   	OWF_Key[313,9]:=1836248757;
   	OWF_Key[313,10]:=799041735;
   	OWF_Key[313,11]:=206920278;
   	OWF_Key[313,12]:=1670185075;
   	OWF_Key[314,0]:=167288513;
   	OWF_Key[314,1]:=1823765264;
   	OWF_Key[314,2]:=1024405687;
   	OWF_Key[314,3]:=1305159346;
   	OWF_Key[314,4]:=1207657799;
   	OWF_Key[314,5]:=1657238232;
   	OWF_Key[314,6]:=1138840138;
   	OWF_Key[314,7]:=1308155371;
   	OWF_Key[314,8]:=444304420;
   	OWF_Key[314,9]:=1715667803;
   	OWF_Key[314,10]:=1632149366;
   	OWF_Key[314,11]:=1040296018;
   	OWF_Key[314,12]:=849669682;
   	OWF_Key[315,0]:=1740950156;
   	OWF_Key[315,1]:=1459336126;
   	OWF_Key[315,2]:=328628267;
   	OWF_Key[315,3]:=1203080453;
   	OWF_Key[315,4]:=244458550;
   	OWF_Key[315,5]:=339011493;
   	OWF_Key[315,6]:=288413275;
   	OWF_Key[315,7]:=1819454890;
   	OWF_Key[315,8]:=1845362003;
   	OWF_Key[315,9]:=298951192;
   	OWF_Key[315,10]:=1589682586;
   	OWF_Key[315,11]:=16248948;
   	OWF_Key[315,12]:=456912391;
   	OWF_Key[316,0]:=1567461601;
   	OWF_Key[316,1]:=1504866295;
   	OWF_Key[316,2]:=356570198;
   	OWF_Key[316,3]:=1868984923;
   	OWF_Key[316,4]:=1342710010;
   	OWF_Key[316,5]:=1358266928;
   	OWF_Key[316,6]:=2133859017;
   	OWF_Key[316,7]:=1343219274;
   	OWF_Key[316,8]:=615300734;
   	OWF_Key[316,9]:=442293248;
   	OWF_Key[316,10]:=115569328;
   	OWF_Key[316,11]:=411515835;
   	OWF_Key[316,12]:=980722739;
   	OWF_Key[317,0]:=1617101216;
   	OWF_Key[317,1]:=1427926010;
   	OWF_Key[317,2]:=1501690115;
   	OWF_Key[317,3]:=1572332995;
   	OWF_Key[317,4]:=766803023;
   	OWF_Key[317,5]:=344781919;
   	OWF_Key[317,6]:=202355058;
   	OWF_Key[317,7]:=1645686166;
   	OWF_Key[317,8]:=2038469782;
   	OWF_Key[317,9]:=932626065;
   	OWF_Key[317,10]:=303846137;
   	OWF_Key[317,11]:=1555884126;
   	OWF_Key[317,12]:=1645831348;
   	OWF_Key[318,0]:=1911130045;
   	OWF_Key[318,1]:=1118008878;
   	OWF_Key[318,2]:=1494023014;
   	OWF_Key[318,3]:=2107585208;
   	OWF_Key[318,4]:=284713769;
   	OWF_Key[318,5]:=1796723039;
   	OWF_Key[318,6]:=1727201322;
   	OWF_Key[318,7]:=1190668856;
   	OWF_Key[318,8]:=1339095212;
   	OWF_Key[318,9]:=173406864;
   	OWF_Key[318,10]:=712994794;
   	OWF_Key[318,11]:=1984462135;
   	OWF_Key[318,12]:=1324617522;
   	OWF_Key[319,0]:=710317526;
   	OWF_Key[319,1]:=2143470138;
   	OWF_Key[319,2]:=1141559794;
   	OWF_Key[319,3]:=1020067858;
   	OWF_Key[319,4]:=1212573818;
   	OWF_Key[319,5]:=251950516;
   	OWF_Key[319,6]:=486915894;
   	OWF_Key[319,7]:=1168168619;
   	OWF_Key[319,8]:=875623503;
   	OWF_Key[319,9]:=1225053274;
   	OWF_Key[319,10]:=1841658760;
   	OWF_Key[319,11]:=643384922;
   	OWF_Key[319,12]:=1498932505;
   	OWF_Key[320,0]:=102598693;
   	OWF_Key[320,1]:=2006227916;
   	OWF_Key[320,2]:=2111704340;
   	OWF_Key[320,3]:=1327817111;
   	OWF_Key[320,4]:=533998976;
   	OWF_Key[320,5]:=682528378;
   	OWF_Key[320,6]:=1146731486;
   	OWF_Key[320,7]:=314830044;
   	OWF_Key[320,8]:=1444899095;
   	OWF_Key[320,9]:=1255844466;
   	OWF_Key[320,10]:=1845456412;
   	OWF_Key[320,11]:=617263051;
   	OWF_Key[320,12]:=1903230993;
   	OWF_Key[321,0]:=728563185;
   	OWF_Key[321,1]:=2118348006;
   	OWF_Key[321,2]:=137733814;
   	OWF_Key[321,3]:=1960321702;
   	OWF_Key[321,4]:=1994024800;
   	OWF_Key[321,5]:=1055124534;
   	OWF_Key[321,6]:=1184942775;
   	OWF_Key[321,7]:=1042106146;
   	OWF_Key[321,8]:=365815672;
   	OWF_Key[321,9]:=482199939;
   	OWF_Key[321,10]:=1674309649;
   	OWF_Key[321,11]:=107218401;
   	OWF_Key[321,12]:=1482710001;
   	OWF_Key[322,0]:=480140151;
   	OWF_Key[322,1]:=1664157226;
   	OWF_Key[322,2]:=1385777309;
   	OWF_Key[322,3]:=1031880165;
   	OWF_Key[322,4]:=1884376959;
   	OWF_Key[322,5]:=816360345;
   	OWF_Key[322,6]:=726566162;
   	OWF_Key[322,7]:=1806503671;
   	OWF_Key[322,8]:=1553960926;
   	OWF_Key[322,9]:=175468279;
   	OWF_Key[322,10]:=851200152;
   	OWF_Key[322,11]:=1218489456;
   	OWF_Key[322,12]:=1327038342;
   	OWF_Key[323,0]:=703604444;
   	OWF_Key[323,1]:=715465034;
   	OWF_Key[323,2]:=1289642010;
   	OWF_Key[323,3]:=699248656;
   	OWF_Key[323,4]:=1691703533;
   	OWF_Key[323,5]:=759781190;
   	OWF_Key[323,6]:=1245758571;
   	OWF_Key[323,7]:=1756157572;
   	OWF_Key[323,8]:=1090534857;
   	OWF_Key[323,9]:=1796279398;
   	OWF_Key[323,10]:=2112880522;
   	OWF_Key[323,11]:=1516054896;
   	OWF_Key[323,12]:=1204227624;
   	OWF_Key[324,0]:=2033719950;
   	OWF_Key[324,1]:=880201031;
   	OWF_Key[324,2]:=1803230991;
   	OWF_Key[324,3]:=621293666;
   	OWF_Key[324,4]:=1059421886;
   	OWF_Key[324,5]:=1417059686;
   	OWF_Key[324,6]:=1107597007;
   	OWF_Key[324,7]:=1754273916;
   	OWF_Key[324,8]:=286719276;
   	OWF_Key[324,9]:=1335157779;
   	OWF_Key[324,10]:=1270792504;
   	OWF_Key[324,11]:=1429366698;
   	OWF_Key[324,12]:=168858728;
   	OWF_Key[325,0]:=1293681434;
   	OWF_Key[325,1]:=1535345076;
   	OWF_Key[325,2]:=1388452763;
   	OWF_Key[325,3]:=55530599;
   	OWF_Key[325,4]:=318445543;
   	OWF_Key[325,5]:=1497513033;
   	OWF_Key[325,6]:=670060474;
   	OWF_Key[325,7]:=406327474;
   	OWF_Key[325,8]:=1513514191;
   	OWF_Key[325,9]:=1367734156;
   	OWF_Key[325,10]:=1652255998;
   	OWF_Key[325,11]:=1424588754;
   	OWF_Key[325,12]:=610648470;
   	OWF_Key[326,0]:=590487839;
   	OWF_Key[326,1]:=1750228599;
   	OWF_Key[326,2]:=894576101;
   	OWF_Key[326,3]:=1294234124;
   	OWF_Key[326,4]:=1878710405;
   	OWF_Key[326,5]:=146757060;
   	OWF_Key[326,6]:=1119600363;
   	OWF_Key[326,7]:=856173152;
   	OWF_Key[326,8]:=1041527179;
   	OWF_Key[326,9]:=362313398;
   	OWF_Key[326,10]:=1714901784;
   	OWF_Key[326,11]:=2028215347;
   	OWF_Key[326,12]:=531940100;
   	OWF_Key[327,0]:=1671026782;
   	OWF_Key[327,1]:=1169850347;
   	OWF_Key[327,2]:=1134426907;
   	OWF_Key[327,3]:=1292812525;
   	OWF_Key[327,4]:=101798530;
   	OWF_Key[327,5]:=1238296398;
   	OWF_Key[327,6]:=306393687;
   	OWF_Key[327,7]:=1147446271;
   	OWF_Key[327,8]:=1224381235;
   	OWF_Key[327,9]:=1992836791;
   	OWF_Key[327,10]:=1945856253;
   	OWF_Key[327,11]:=1597999087;
   	OWF_Key[327,12]:=805381885;
   	OWF_Key[328,0]:=202644485;
   	OWF_Key[328,1]:=1993247;
   	OWF_Key[328,2]:=1069190287;
   	OWF_Key[328,3]:=36265956;
   	OWF_Key[328,4]:=984589841;
   	OWF_Key[328,5]:=1964325587;
   	OWF_Key[328,6]:=1822401321;
   	OWF_Key[328,7]:=1581068640;
   	OWF_Key[328,8]:=1946895186;
   	OWF_Key[328,9]:=1040124109;
   	OWF_Key[328,10]:=177594935;
   	OWF_Key[328,11]:=810665212;
   	OWF_Key[328,12]:=538300843;
   	OWF_Key[329,0]:=358177491;
   	OWF_Key[329,1]:=14270137;
   	OWF_Key[329,2]:=1493093187;
   	OWF_Key[329,3]:=919469069;
   	OWF_Key[329,4]:=1050322522;
   	OWF_Key[329,5]:=777998955;
   	OWF_Key[329,6]:=575835217;
   	OWF_Key[329,7]:=734728415;
   	OWF_Key[329,8]:=1687372136;
   	OWF_Key[329,9]:=120770498;
   	OWF_Key[329,10]:=234291522;
   	OWF_Key[329,11]:=1039125923;
   	OWF_Key[329,12]:=416355858;
   	OWF_Key[330,0]:=1943253149;
   	OWF_Key[330,1]:=1471630074;
   	OWF_Key[330,2]:=216018934;
   	OWF_Key[330,3]:=1374893637;
   	OWF_Key[330,4]:=1074805829;
   	OWF_Key[330,5]:=372858553;
   	OWF_Key[330,6]:=1175946170;
   	OWF_Key[330,7]:=858540876;
   	OWF_Key[330,8]:=1753558902;
   	OWF_Key[330,9]:=1707867970;
   	OWF_Key[330,10]:=1046672431;
   	OWF_Key[330,11]:=321627573;
   	OWF_Key[330,12]:=953995245;
   	OWF_Key[331,0]:=189455458;
   	OWF_Key[331,1]:=1009326955;
   	OWF_Key[331,2]:=1832939834;
   	OWF_Key[331,3]:=2134573027;
   	OWF_Key[331,4]:=87610150;
   	OWF_Key[331,5]:=1728917062;
   	OWF_Key[331,6]:=431488573;
   	OWF_Key[331,7]:=1128489670;
   	OWF_Key[331,8]:=2097887200;
   	OWF_Key[331,9]:=648619132;
   	OWF_Key[331,10]:=1706988526;
   	OWF_Key[331,11]:=726343804;
   	OWF_Key[331,12]:=707324238;
   	OWF_Key[332,0]:=991909150;
   	OWF_Key[332,1]:=241527182;
   	OWF_Key[332,2]:=1117912615;
   	OWF_Key[332,3]:=1742565370;
   	OWF_Key[332,4]:=847260552;
   	OWF_Key[332,5]:=695992848;
   	OWF_Key[332,6]:=2124266459;
   	OWF_Key[332,7]:=3760078;
   	OWF_Key[332,8]:=1788157085;
   	OWF_Key[332,9]:=311304058;
   	OWF_Key[332,10]:=881662921;
   	OWF_Key[332,11]:=1394957333;
   	OWF_Key[332,12]:=1120352024;
   	OWF_Key[333,0]:=2017580647;
   	OWF_Key[333,1]:=1876652258;
   	OWF_Key[333,2]:=764862997;
   	OWF_Key[333,3]:=880722372;
   	OWF_Key[333,4]:=552911306;
   	OWF_Key[333,5]:=246790094;
   	OWF_Key[333,6]:=24871650;
   	OWF_Key[333,7]:=1141621677;
   	OWF_Key[333,8]:=901566941;
   	OWF_Key[333,9]:=1841434757;
   	OWF_Key[333,10]:=1041061206;
   	OWF_Key[333,11]:=1725521277;
   	OWF_Key[333,12]:=215989094;
   	OWF_Key[334,0]:=1359582125;
   	OWF_Key[334,1]:=1101587530;
   	OWF_Key[334,2]:=643671334;
   	OWF_Key[334,3]:=182418752;
   	OWF_Key[334,4]:=90220878;
   	OWF_Key[334,5]:=1699068097;
   	OWF_Key[334,6]:=2002200371;
   	OWF_Key[334,7]:=636677458;
   	OWF_Key[334,8]:=1791268416;
   	OWF_Key[334,9]:=675643818;
   	OWF_Key[334,10]:=503721560;
   	OWF_Key[334,11]:=510726541;
   	OWF_Key[334,12]:=1493156750;
   	OWF_Key[335,0]:=2104270054;
   	OWF_Key[335,1]:=1342954771;
   	OWF_Key[335,2]:=383320059;
   	OWF_Key[335,3]:=32507010;
   	OWF_Key[335,4]:=145617757;
   	OWF_Key[335,5]:=2071263462;
   	OWF_Key[335,6]:=418578355;
   	OWF_Key[335,7]:=1568019122;
   	OWF_Key[335,8]:=1378841819;
   	OWF_Key[335,9]:=881582072;
   	OWF_Key[335,10]:=451327839;
   	OWF_Key[335,11]:=392128201;
   	OWF_Key[335,12]:=2080483153;
   	OWF_Key[336,0]:=1121801471;
   	OWF_Key[336,1]:=181935598;
   	OWF_Key[336,2]:=1577536789;
   	OWF_Key[336,3]:=338027538;
   	OWF_Key[336,4]:=373853370;
   	OWF_Key[336,5]:=426935573;
   	OWF_Key[336,6]:=452734870;
   	OWF_Key[336,7]:=652861449;
   	OWF_Key[336,8]:=139824699;
   	OWF_Key[336,9]:=1109137398;
   	OWF_Key[336,10]:=858218833;
   	OWF_Key[336,11]:=479988425;
   	OWF_Key[336,12]:=1896055883;
   	OWF_Key[337,0]:=568312635;
   	OWF_Key[337,1]:=1548749383;
   	OWF_Key[337,2]:=1997225580;
   	OWF_Key[337,3]:=1096216702;
   	OWF_Key[337,4]:=1224318064;
   	OWF_Key[337,5]:=616115760;
   	OWF_Key[337,6]:=291003252;
   	OWF_Key[337,7]:=1233051881;
   	OWF_Key[337,8]:=504389448;
   	OWF_Key[337,9]:=318158703;
   	OWF_Key[337,10]:=1063373500;
   	OWF_Key[337,11]:=91958396;
   	OWF_Key[337,12]:=1275563904;
   	OWF_Key[338,0]:=1517460097;
   	OWF_Key[338,1]:=646770227;
   	OWF_Key[338,2]:=1122144401;
   	OWF_Key[338,3]:=565403386;
   	OWF_Key[338,4]:=1212489744;
   	OWF_Key[338,5]:=1998449907;
   	OWF_Key[338,6]:=1155005407;
   	OWF_Key[338,7]:=1204471807;
   	OWF_Key[338,8]:=629732107;
   	OWF_Key[338,9]:=436852736;
   	OWF_Key[338,10]:=399692315;
   	OWF_Key[338,11]:=46670747;
   	OWF_Key[338,12]:=651743739;
   	OWF_Key[339,0]:=411731057;
   	OWF_Key[339,1]:=1025513189;
   	OWF_Key[339,2]:=682007003;
   	OWF_Key[339,3]:=148663973;
   	OWF_Key[339,4]:=568231694;
   	OWF_Key[339,5]:=475104531;
   	OWF_Key[339,6]:=1114405893;
   	OWF_Key[339,7]:=1730439593;
   	OWF_Key[339,8]:=1646413011;
   	OWF_Key[339,9]:=1222983612;
   	OWF_Key[339,10]:=1114304189;
   	OWF_Key[339,11]:=1118366461;
   	OWF_Key[339,12]:=585111365;
   	OWF_Key[340,0]:=101941386;
   	OWF_Key[340,1]:=91975525;
   	OWF_Key[340,2]:=935751465;
   	OWF_Key[340,3]:=1019109662;
   	OWF_Key[340,4]:=1672840690;
   	OWF_Key[340,5]:=1717134215;
   	OWF_Key[340,6]:=582105036;
   	OWF_Key[340,7]:=2001867664;
   	OWF_Key[340,8]:=1828725794;
   	OWF_Key[340,9]:=295780255;
   	OWF_Key[340,10]:=226565605;
   	OWF_Key[340,11]:=140644531;
   	OWF_Key[340,12]:=955234534;
   	OWF_Key[341,0]:=101214910;
   	OWF_Key[341,1]:=1797184804;
   	OWF_Key[341,2]:=1590624389;
   	OWF_Key[341,3]:=274218088;
   	OWF_Key[341,4]:=1400290409;
   	OWF_Key[341,5]:=622516308;
   	OWF_Key[341,6]:=266931326;
   	OWF_Key[341,7]:=1008039898;
   	OWF_Key[341,8]:=349311417;
   	OWF_Key[341,9]:=98462939;
   	OWF_Key[341,10]:=1692269881;
   	OWF_Key[341,11]:=335797834;
   	OWF_Key[341,12]:=1907594453;
   	OWF_Key[342,0]:=1231887310;
   	OWF_Key[342,1]:=1325769248;
   	OWF_Key[342,2]:=2004054930;
   	OWF_Key[342,3]:=279890262;
   	OWF_Key[342,4]:=361598874;
   	OWF_Key[342,5]:=1171465859;
   	OWF_Key[342,6]:=2070486323;
   	OWF_Key[342,7]:=1882949837;
   	OWF_Key[342,8]:=953594315;
   	OWF_Key[342,9]:=14687673;
   	OWF_Key[342,10]:=270943799;
   	OWF_Key[342,11]:=214886758;
   	OWF_Key[342,12]:=558480261;
   	OWF_Key[343,0]:=1964622833;
   	OWF_Key[343,1]:=1098443067;
   	OWF_Key[343,2]:=812239160;
   	OWF_Key[343,3]:=587893861;
   	OWF_Key[343,4]:=967632277;
   	OWF_Key[343,5]:=1068169670;
   	OWF_Key[343,6]:=227120408;
   	OWF_Key[343,7]:=1873201141;
   	OWF_Key[343,8]:=2035351652;
   	OWF_Key[343,9]:=1498518442;
   	OWF_Key[343,10]:=22841995;
   	OWF_Key[343,11]:=858808412;
   	OWF_Key[343,12]:=1607329516;
   	OWF_Key[344,0]:=1130671788;
   	OWF_Key[344,1]:=1611076207;
   	OWF_Key[344,2]:=242483588;
   	OWF_Key[344,3]:=809041729;
   	OWF_Key[344,4]:=400295578;
   	OWF_Key[344,5]:=2143399394;
   	OWF_Key[344,6]:=58120252;
   	OWF_Key[344,7]:=1105914141;
   	OWF_Key[344,8]:=65538387;
   	OWF_Key[344,9]:=1432524579;
   	OWF_Key[344,10]:=1081012900;
   	OWF_Key[344,11]:=55469365;
   	OWF_Key[344,12]:=309634431;
   	OWF_Key[345,0]:=684582410;
   	OWF_Key[345,1]:=1095651926;
   	OWF_Key[345,2]:=153896313;
   	OWF_Key[345,3]:=822841261;
   	OWF_Key[345,4]:=1221560818;
   	OWF_Key[345,5]:=1231028825;
   	OWF_Key[345,6]:=897926319;
   	OWF_Key[345,7]:=1460520646;
   	OWF_Key[345,8]:=1889402372;
   	OWF_Key[345,9]:=924838793;
   	OWF_Key[345,10]:=89408900;
   	OWF_Key[345,11]:=14556754;
   	OWF_Key[345,12]:=1730121170;
   	OWF_Key[346,0]:=1005743598;
   	OWF_Key[346,1]:=1774083544;
   	OWF_Key[346,2]:=825020351;
   	OWF_Key[346,3]:=1019981492;
   	OWF_Key[346,4]:=1125356371;
   	OWF_Key[346,5]:=1083900510;
   	OWF_Key[346,6]:=1609438256;
   	OWF_Key[346,7]:=540419995;
   	OWF_Key[346,8]:=1053298608;
   	OWF_Key[346,9]:=1871567025;
   	OWF_Key[346,10]:=279687974;
   	OWF_Key[346,11]:=1659531677;
   	OWF_Key[346,12]:=893635376;
   	OWF_Key[347,0]:=1555577303;
   	OWF_Key[347,1]:=1413413491;
   	OWF_Key[347,2]:=2095683958;
   	OWF_Key[347,3]:=4648522;
   	OWF_Key[347,4]:=810466289;
   	OWF_Key[347,5]:=645762303;
   	OWF_Key[347,6]:=1915839225;
   	OWF_Key[347,7]:=1204668640;
   	OWF_Key[347,8]:=368397103;
   	OWF_Key[347,9]:=1534490663;
   	OWF_Key[347,10]:=1060404450;
   	OWF_Key[347,11]:=1757654932;
   	OWF_Key[347,12]:=1194908497;
   	OWF_Key[348,0]:=1516532639;
   	OWF_Key[348,1]:=2013259281;
   	OWF_Key[348,2]:=2061450127;
   	OWF_Key[348,3]:=1191764982;
   	OWF_Key[348,4]:=1951391276;
   	OWF_Key[348,5]:=269341694;
   	OWF_Key[348,6]:=1635172496;
   	OWF_Key[348,7]:=380270759;
   	OWF_Key[348,8]:=1409414929;
   	OWF_Key[348,9]:=247162533;
   	OWF_Key[348,10]:=1466424841;
   	OWF_Key[348,11]:=151341368;
   	OWF_Key[348,12]:=1022982709;
   	OWF_Key[349,0]:=943486149;
   	OWF_Key[349,1]:=1407267179;
   	OWF_Key[349,2]:=669896272;
   	OWF_Key[349,3]:=1384608088;
   	OWF_Key[349,4]:=1373845006;
   	OWF_Key[349,5]:=283357154;
   	OWF_Key[349,6]:=1997522781;
   	OWF_Key[349,7]:=1432204524;
   	OWF_Key[349,8]:=1952512283;
   	OWF_Key[349,9]:=917951409;
   	OWF_Key[349,10]:=1175316246;
   	OWF_Key[349,11]:=1303327261;
   	OWF_Key[349,12]:=993699275;
   	OWF_Key[350,0]:=200790839;
   	OWF_Key[350,1]:=1254080954;
   	OWF_Key[350,2]:=269083328;
   	OWF_Key[350,3]:=451236702;
   	OWF_Key[350,4]:=1810271156;
   	OWF_Key[350,5]:=398842525;
   	OWF_Key[350,6]:=2045546455;
   	OWF_Key[350,7]:=1383822173;
   	OWF_Key[350,8]:=165988296;
   	OWF_Key[350,9]:=178683914;
   	OWF_Key[350,10]:=1579074927;
   	OWF_Key[350,11]:=2038230152;
   	OWF_Key[350,12]:=1948721857;
   	OWF_Key[351,0]:=195262027;
   	OWF_Key[351,1]:=654194628;
   	OWF_Key[351,2]:=1538814138;
   	OWF_Key[351,3]:=754899861;
   	OWF_Key[351,4]:=1491407397;
   	OWF_Key[351,5]:=2144262794;
   	OWF_Key[351,6]:=2081529130;
   	OWF_Key[351,7]:=237406198;
   	OWF_Key[351,8]:=730746525;
   	OWF_Key[351,9]:=45813349;
   	OWF_Key[351,10]:=772554456;
   	OWF_Key[351,11]:=1135823331;
   	OWF_Key[351,12]:=1908013618;
   	OWF_Key[352,0]:=629896472;
   	OWF_Key[352,1]:=959658323;
   	OWF_Key[352,2]:=271563843;
   	OWF_Key[352,3]:=151103786;
   	OWF_Key[352,4]:=198227326;
   	OWF_Key[352,5]:=1503636945;
   	OWF_Key[352,6]:=1183422528;
   	OWF_Key[352,7]:=63370702;
   	OWF_Key[352,8]:=676432682;
   	OWF_Key[352,9]:=547620457;
   	OWF_Key[352,10]:=47116289;
   	OWF_Key[352,11]:=439158043;
   	OWF_Key[352,12]:=360603174;
   	OWF_Key[353,0]:=1822681441;
   	OWF_Key[353,1]:=954624633;
   	OWF_Key[353,2]:=1755380528;
   	OWF_Key[353,3]:=487961148;
   	OWF_Key[353,4]:=259695196;
   	OWF_Key[353,5]:=509804854;
   	OWF_Key[353,6]:=252112419;
   	OWF_Key[353,7]:=983541593;
   	OWF_Key[353,8]:=1268917091;
   	OWF_Key[353,9]:=257094738;
   	OWF_Key[353,10]:=247380732;
   	OWF_Key[353,11]:=65856510;
   	OWF_Key[353,12]:=906386107;
   	OWF_Key[354,0]:=1743785763;
   	OWF_Key[354,1]:=550061803;
   	OWF_Key[354,2]:=285850847;
   	OWF_Key[354,3]:=296303136;
   	OWF_Key[354,4]:=637258478;
   	OWF_Key[354,5]:=995436917;
   	OWF_Key[354,6]:=934855509;
   	OWF_Key[354,7]:=805099594;
   	OWF_Key[354,8]:=830609290;
   	OWF_Key[354,9]:=1989592865;
   	OWF_Key[354,10]:=770381295;
   	OWF_Key[354,11]:=85185801;
   	OWF_Key[354,12]:=1089481680;
   	OWF_Key[355,0]:=335583696;
   	OWF_Key[355,1]:=1301561535;
   	OWF_Key[355,2]:=1154445123;
   	OWF_Key[355,3]:=1382772528;
   	OWF_Key[355,4]:=1524115461;
   	OWF_Key[355,5]:=699342829;
   	OWF_Key[355,6]:=405837931;
   	OWF_Key[355,7]:=114037572;
   	OWF_Key[355,8]:=439771994;
   	OWF_Key[355,9]:=486638158;
   	OWF_Key[355,10]:=1997470365;
   	OWF_Key[355,11]:=1883749861;
   	OWF_Key[355,12]:=1382653884;
   	OWF_Key[356,0]:=1115691661;
   	OWF_Key[356,1]:=258797628;
   	OWF_Key[356,2]:=93806010;
   	OWF_Key[356,3]:=1280185665;
   	OWF_Key[356,4]:=1365529581;
   	OWF_Key[356,5]:=1561953534;
   	OWF_Key[356,6]:=904506324;
   	OWF_Key[356,7]:=1353500892;
   	OWF_Key[356,8]:=2131662628;
   	OWF_Key[356,9]:=1593427382;
   	OWF_Key[356,10]:=387540744;
   	OWF_Key[356,11]:=744268773;
   	OWF_Key[356,12]:=519696264;
   	OWF_Key[357,0]:=1578539292;
   	OWF_Key[357,1]:=562385808;
   	OWF_Key[357,2]:=613815707;
   	OWF_Key[357,3]:=111408283;
   	OWF_Key[357,4]:=822552011;
   	OWF_Key[357,5]:=1056326650;
   	OWF_Key[357,6]:=1089048739;
   	OWF_Key[357,7]:=1236032568;
   	OWF_Key[357,8]:=899502552;
   	OWF_Key[357,9]:=293770547;
   	OWF_Key[357,10]:=1802477383;
   	OWF_Key[357,11]:=432228269;
   	OWF_Key[357,12]:=1447757393;
   	OWF_Key[358,0]:=1730852905;
   	OWF_Key[358,1]:=784052714;
   	OWF_Key[358,2]:=1551124257;
   	OWF_Key[358,3]:=850463373;
   	OWF_Key[358,4]:=613821989;
   	OWF_Key[358,5]:=558345880;
   	OWF_Key[358,6]:=485866837;
   	OWF_Key[358,7]:=747598701;
   	OWF_Key[358,8]:=175180911;
   	OWF_Key[358,9]:=1874092731;
   	OWF_Key[358,10]:=465240862;
   	OWF_Key[358,11]:=1166967805;
   	OWF_Key[358,12]:=606152266;
   	OWF_Key[359,0]:=900648406;
   	OWF_Key[359,1]:=2075197520;
   	OWF_Key[359,2]:=108720043;
   	OWF_Key[359,3]:=1645648917;
   	OWF_Key[359,4]:=568308072;
   	OWF_Key[359,5]:=742876145;
   	OWF_Key[359,6]:=287513467;
   	OWF_Key[359,7]:=545461664;
   	OWF_Key[359,8]:=726036885;
   	OWF_Key[359,9]:=1357184276;
   	OWF_Key[359,10]:=1587129830;
   	OWF_Key[359,11]:=920264815;
   	OWF_Key[359,12]:=1013402406;
   	OWF_Key[360,0]:=177604624;
   	OWF_Key[360,1]:=32739705;
   	OWF_Key[360,2]:=2072866395;
   	OWF_Key[360,3]:=924854198;
   	OWF_Key[360,4]:=102148350;
   	OWF_Key[360,5]:=624243173;
   	OWF_Key[360,6]:=1547779740;
   	OWF_Key[360,7]:=769169699;
   	OWF_Key[360,8]:=1606576629;
   	OWF_Key[360,9]:=642360978;
   	OWF_Key[360,10]:=162193754;
   	OWF_Key[360,11]:=826106027;
   	OWF_Key[360,12]:=30502231;
   	OWF_Key[361,0]:=1256538179;
   	OWF_Key[361,1]:=141218112;
   	OWF_Key[361,2]:=751607397;
   	OWF_Key[361,3]:=1908899164;
   	OWF_Key[361,4]:=646341656;
   	OWF_Key[361,5]:=1891616426;
   	OWF_Key[361,6]:=365239531;
   	OWF_Key[361,7]:=1574850028;
   	OWF_Key[361,8]:=1988244313;
   	OWF_Key[361,9]:=1740473693;
   	OWF_Key[361,10]:=802008055;
   	OWF_Key[361,11]:=126991285;
   	OWF_Key[361,12]:=28306954;
   	OWF_Key[362,0]:=131619368;
   	OWF_Key[362,1]:=2007697757;
   	OWF_Key[362,2]:=1655931393;
   	OWF_Key[362,3]:=1047467215;
   	OWF_Key[362,4]:=1636337202;
   	OWF_Key[362,5]:=472117744;
   	OWF_Key[362,6]:=1508581209;
   	OWF_Key[362,7]:=621372235;
   	OWF_Key[362,8]:=523575959;
   	OWF_Key[362,9]:=1226782044;
   	OWF_Key[362,10]:=1900906814;
   	OWF_Key[362,11]:=1885885148;
   	OWF_Key[362,12]:=1461350739;
   	OWF_Key[363,0]:=1096238794;
   	OWF_Key[363,1]:=2100318410;
   	OWF_Key[363,2]:=335439393;
   	OWF_Key[363,3]:=1020314535;
   	OWF_Key[363,4]:=1221649134;
   	OWF_Key[363,5]:=226531355;
   	OWF_Key[363,6]:=2050792586;
   	OWF_Key[363,7]:=1825771681;
   	OWF_Key[363,8]:=622633333;
   	OWF_Key[363,9]:=539910382;
   	OWF_Key[363,10]:=331725508;
   	OWF_Key[363,11]:=1362579679;
   	OWF_Key[363,12]:=659996391;
   	OWF_Key[364,0]:=1223229109;
   	OWF_Key[364,1]:=2092484739;
   	OWF_Key[364,2]:=1264224138;
   	OWF_Key[364,3]:=570346107;
   	OWF_Key[364,4]:=1964626207;
   	OWF_Key[364,5]:=1408734319;
   	OWF_Key[364,6]:=1845742860;
   	OWF_Key[364,7]:=402751573;
   	OWF_Key[364,8]:=1939948710;
   	OWF_Key[364,9]:=1584034187;
   	OWF_Key[364,10]:=595028108;
   	OWF_Key[364,11]:=1414436209;
   	OWF_Key[364,12]:=1847538317;
   	OWF_Key[365,0]:=4015651;
   	OWF_Key[365,1]:=1160278100;
   	OWF_Key[365,2]:=2133678767;
   	OWF_Key[365,3]:=711727851;
   	OWF_Key[365,4]:=767763311;
   	OWF_Key[365,5]:=1454993297;
   	OWF_Key[365,6]:=1460694151;
   	OWF_Key[365,7]:=525797765;
   	OWF_Key[365,8]:=850336057;
   	OWF_Key[365,9]:=1219415484;
   	OWF_Key[365,10]:=1108439294;
   	OWF_Key[365,11]:=1902590331;
   	OWF_Key[365,12]:=906794746;
   	OWF_Key[366,0]:=403671914;
   	OWF_Key[366,1]:=1058773782;
   	OWF_Key[366,2]:=1656204258;
   	OWF_Key[366,3]:=1592499955;
   	OWF_Key[366,4]:=49767413;
   	OWF_Key[366,5]:=409347063;
   	OWF_Key[366,6]:=1649695713;
   	OWF_Key[366,7]:=158765815;
   	OWF_Key[366,8]:=1095400275;
   	OWF_Key[366,9]:=940994704;
   	OWF_Key[366,10]:=108034986;
   	OWF_Key[366,11]:=752356231;
   	OWF_Key[366,12]:=814289094;
   	OWF_Key[367,0]:=893533826;
   	OWF_Key[367,1]:=1017742775;
   	OWF_Key[367,2]:=1388320011;
   	OWF_Key[367,3]:=1380629462;
   	OWF_Key[367,4]:=1569037800;
   	OWF_Key[367,5]:=914194369;
   	OWF_Key[367,6]:=1663813751;
   	OWF_Key[367,7]:=1583027395;
   	OWF_Key[367,8]:=1218601859;
   	OWF_Key[367,9]:=720386169;
   	OWF_Key[367,10]:=219130365;
   	OWF_Key[367,11]:=784479652;
   	OWF_Key[367,12]:=555792365;
   	OWF_Key[368,0]:=325492182;
   	OWF_Key[368,1]:=1070949215;
   	OWF_Key[368,2]:=1612439119;
   	OWF_Key[368,3]:=520339558;
   	OWF_Key[368,4]:=283026555;
   	OWF_Key[368,5]:=397262156;
   	OWF_Key[368,6]:=1543948565;
   	OWF_Key[368,7]:=1944054940;
   	OWF_Key[368,8]:=1555674573;
   	OWF_Key[368,9]:=602776568;
   	OWF_Key[368,10]:=427610564;
   	OWF_Key[368,11]:=839181682;
   	OWF_Key[368,12]:=580284637;
   	OWF_Key[369,0]:=1845577166;
   	OWF_Key[369,1]:=755980584;
   	OWF_Key[369,2]:=1870933655;
   	OWF_Key[369,3]:=1185025747;
   	OWF_Key[369,4]:=966601097;
   	OWF_Key[369,5]:=1097318171;
   	OWF_Key[369,6]:=670129362;
   	OWF_Key[369,7]:=584817892;
   	OWF_Key[369,8]:=1165106007;
   	OWF_Key[369,9]:=1620962611;
   	OWF_Key[369,10]:=357961287;
   	OWF_Key[369,11]:=861787749;
   	OWF_Key[369,12]:=241787703;
   	OWF_Key[370,0]:=942018444;
   	OWF_Key[370,1]:=1269279705;
   	OWF_Key[370,2]:=1263220557;
   	OWF_Key[370,3]:=1356082571;
   	OWF_Key[370,4]:=1113501611;
   	OWF_Key[370,5]:=901687732;
   	OWF_Key[370,6]:=724787856;
   	OWF_Key[370,7]:=1857871907;
   	OWF_Key[370,8]:=1656844551;
   	OWF_Key[370,9]:=306802645;
   	OWF_Key[370,10]:=2100992171;
   	OWF_Key[370,11]:=52296823;
   	OWF_Key[370,12]:=902420557;
   	OWF_Key[371,0]:=1269415789;
   	OWF_Key[371,1]:=2005771722;
   	OWF_Key[371,2]:=586171040;
   	OWF_Key[371,3]:=165451393;
   	OWF_Key[371,4]:=576615512;
   	OWF_Key[371,5]:=527546538;
   	OWF_Key[371,6]:=1303775377;
   	OWF_Key[371,7]:=521781338;
   	OWF_Key[371,8]:=1537585392;
   	OWF_Key[371,9]:=78099681;
   	OWF_Key[371,10]:=67338240;
   	OWF_Key[371,11]:=602320789;
   	OWF_Key[371,12]:=1337869044;
   	OWF_Key[372,0]:=227580228;
   	OWF_Key[372,1]:=329197407;
   	OWF_Key[372,2]:=572336303;
   	OWF_Key[372,3]:=170847879;
   	OWF_Key[372,4]:=1928684315;
   	OWF_Key[372,5]:=1482343427;
   	OWF_Key[372,6]:=1503790864;
   	OWF_Key[372,7]:=978039587;
   	OWF_Key[372,8]:=96787721;
   	OWF_Key[372,9]:=1634589016;
   	OWF_Key[372,10]:=887352446;
   	OWF_Key[372,11]:=1225710675;
   	OWF_Key[372,12]:=1255583127;
   	OWF_Key[373,0]:=1574805053;
   	OWF_Key[373,1]:=1906524970;
   	OWF_Key[373,2]:=1220831147;
   	OWF_Key[373,3]:=1755035379;
   	OWF_Key[373,4]:=700601326;
   	OWF_Key[373,5]:=116735923;
   	OWF_Key[373,6]:=2112340640;
   	OWF_Key[373,7]:=371913440;
   	OWF_Key[373,8]:=40799741;
   	OWF_Key[373,9]:=947146791;
   	OWF_Key[373,10]:=471104621;
   	OWF_Key[373,11]:=1412203619;
   	OWF_Key[373,12]:=845996704;
   	OWF_Key[374,0]:=428759036;
   	OWF_Key[374,1]:=1624793299;
   	OWF_Key[374,2]:=1944579770;
   	OWF_Key[374,3]:=1792346547;
   	OWF_Key[374,4]:=2140766573;
   	OWF_Key[374,5]:=1878116227;
   	OWF_Key[374,6]:=557805278;
   	OWF_Key[374,7]:=1528393183;
   	OWF_Key[374,8]:=146799061;
   	OWF_Key[374,9]:=1630448555;
   	OWF_Key[374,10]:=1664880067;
   	OWF_Key[374,11]:=1400822156;
   	OWF_Key[374,12]:=1781564781;
   	OWF_Key[375,0]:=1834227907;
   	OWF_Key[375,1]:=1876025053;
   	OWF_Key[375,2]:=403950487;
   	OWF_Key[375,3]:=1869177872;
   	OWF_Key[375,4]:=960241097;
   	OWF_Key[375,5]:=1522005120;
   	OWF_Key[375,6]:=1831743326;
   	OWF_Key[375,7]:=101149434;
   	OWF_Key[375,8]:=375981746;
   	OWF_Key[375,9]:=412110870;
   	OWF_Key[375,10]:=72672528;
   	OWF_Key[375,11]:=1135232175;
   	OWF_Key[375,12]:=1862200496;
   	OWF_Key[376,0]:=1238973653;
   	OWF_Key[376,1]:=864504014;
   	OWF_Key[376,2]:=1385128927;
   	OWF_Key[376,3]:=798071796;
   	OWF_Key[376,4]:=1597649644;
   	OWF_Key[376,5]:=2104447674;
   	OWF_Key[376,6]:=100897745;
   	OWF_Key[376,7]:=538205605;
   	OWF_Key[376,8]:=558079957;
   	OWF_Key[376,9]:=1188859919;
   	OWF_Key[376,10]:=1574973441;
   	OWF_Key[376,11]:=1416257780;
   	OWF_Key[376,12]:=1826775749;
   	OWF_Key[377,0]:=1154584260;
   	OWF_Key[377,1]:=1299724199;
   	OWF_Key[377,2]:=1287894970;
   	OWF_Key[377,3]:=1990190052;
   	OWF_Key[377,4]:=1144015219;
   	OWF_Key[377,5]:=2075114646;
   	OWF_Key[377,6]:=767757119;
   	OWF_Key[377,7]:=1800023041;
   	OWF_Key[377,8]:=1709123131;
   	OWF_Key[377,9]:=980766873;
   	OWF_Key[377,10]:=818219643;
   	OWF_Key[377,11]:=942098504;
   	OWF_Key[377,12]:=1390689164;
   	OWF_Key[378,0]:=746390694;
   	OWF_Key[378,1]:=393623812;
   	OWF_Key[378,2]:=1164801535;
   	OWF_Key[378,3]:=2091357433;
   	OWF_Key[378,4]:=157745671;
   	OWF_Key[378,5]:=863722553;
   	OWF_Key[378,6]:=1525069691;
   	OWF_Key[378,7]:=755533550;
   	OWF_Key[378,8]:=179632376;
   	OWF_Key[378,9]:=449419476;
   	OWF_Key[378,10]:=839028966;
   	OWF_Key[378,11]:=1054098079;
   	OWF_Key[378,12]:=82253776;
   	OWF_Key[379,0]:=1529647443;
   	OWF_Key[379,1]:=1737062437;
   	OWF_Key[379,2]:=857081988;
   	OWF_Key[379,3]:=937415973;
   	OWF_Key[379,4]:=948568225;
   	OWF_Key[379,5]:=789887072;
   	OWF_Key[379,6]:=1084648100;
   	OWF_Key[379,7]:=3197571;
   	OWF_Key[379,8]:=1571124900;
   	OWF_Key[379,9]:=1917543500;
   	OWF_Key[379,10]:=1019946534;
   	OWF_Key[379,11]:=1818027515;
   	OWF_Key[379,12]:=476331063;
   	OWF_Key[380,0]:=1798466443;
   	OWF_Key[380,1]:=2068248887;
   	OWF_Key[380,2]:=361438599;
   	OWF_Key[380,3]:=1090863320;
   	OWF_Key[380,4]:=417076587;
   	OWF_Key[380,5]:=1967089161;
   	OWF_Key[380,6]:=880082427;
   	OWF_Key[380,7]:=1951088809;
   	OWF_Key[380,8]:=1431072;
   	OWF_Key[380,9]:=1223741584;
   	OWF_Key[380,10]:=511310210;
   	OWF_Key[380,11]:=1823630479;
   	OWF_Key[380,12]:=1993212374;
   	OWF_Key[381,0]:=1243769354;
   	OWF_Key[381,1]:=1629593806;
   	OWF_Key[381,2]:=2100292201;
   	OWF_Key[381,3]:=1208010661;
   	OWF_Key[381,4]:=106616940;
   	OWF_Key[381,5]:=962719993;
   	OWF_Key[381,6]:=1154410983;
   	OWF_Key[381,7]:=1870961384;
   	OWF_Key[381,8]:=1052655094;
   	OWF_Key[381,9]:=1225437253;
   	OWF_Key[381,10]:=1199010231;
   	OWF_Key[381,11]:=1619648686;
   	OWF_Key[381,12]:=787437959;
   	OWF_Key[382,0]:=1168123735;
   	OWF_Key[382,1]:=1045160339;
   	OWF_Key[382,2]:=672470685;
   	OWF_Key[382,3]:=1791276252;
   	OWF_Key[382,4]:=1042435383;
   	OWF_Key[382,5]:=768535115;
   	OWF_Key[382,6]:=683097434;
   	OWF_Key[382,7]:=687378611;
   	OWF_Key[382,8]:=1313788124;
   	OWF_Key[382,9]:=802668805;
   	OWF_Key[382,10]:=598443602;
   	OWF_Key[382,11]:=1162520547;
   	OWF_Key[382,12]:=844158402;
   	OWF_Key[383,0]:=91416782;
   	OWF_Key[383,1]:=1237800742;
   	OWF_Key[383,2]:=1669273560;
   	OWF_Key[383,3]:=276647066;
   	OWF_Key[383,4]:=34857035;
   	OWF_Key[383,5]:=996826804;
   	OWF_Key[383,6]:=39317912;
   	OWF_Key[383,7]:=773423270;
   	OWF_Key[383,8]:=15915813;
   	OWF_Key[383,9]:=240056791;
   	OWF_Key[383,10]:=312842243;
   	OWF_Key[383,11]:=1562137978;
   	OWF_Key[383,12]:=289842865;
   End_If;
   If OWF_Ver = 2 Then
   	OWF_Key[0,13]:=134993119;
   	OWF_Key[0,14]:=618806328;
   	OWF_Key[0,15]:=1709154388;
   	OWF_Key[0,16]:=1312484224;
   	OWF_Key[1,13]:=710355550;
   	OWF_Key[1,14]:=1510353068;
   	OWF_Key[1,15]:=2109589066;
   	OWF_Key[1,16]:=1309621689;
   	OWF_Key[2,13]:=1228128301;
   	OWF_Key[2,14]:=709628399;
   	OWF_Key[2,15]:=220820696;
   	OWF_Key[2,16]:=855501000;
   	OWF_Key[3,13]:=1041338116;
   	OWF_Key[3,14]:=626869115;
   	OWF_Key[3,15]:=545726397;
   	OWF_Key[3,16]:=2001122690;
   	OWF_Key[4,13]:=414740093;
   	OWF_Key[4,14]:=333230235;
   	OWF_Key[4,15]:=726355073;
   	OWF_Key[4,16]:=1347715235;
   	OWF_Key[5,13]:=578488929;
   	OWF_Key[5,14]:=356206792;
   	OWF_Key[5,15]:=615836757;
   	OWF_Key[5,16]:=1759694649;
   	OWF_Key[6,13]:=548059399;
   	OWF_Key[6,14]:=2136311382;
   	OWF_Key[6,15]:=1467296399;
   	OWF_Key[6,16]:=293140255;
   	OWF_Key[7,13]:=792442081;
   	OWF_Key[7,14]:=1655991506;
   	OWF_Key[7,15]:=1524245270;
   	OWF_Key[7,16]:=492106621;
   	OWF_Key[8,13]:=1444124688;
   	OWF_Key[8,14]:=2019737066;
   	OWF_Key[8,15]:=562887751;
   	OWF_Key[8,16]:=920287799;
   	OWF_Key[9,13]:=403848183;
   	OWF_Key[9,14]:=405587786;
   	OWF_Key[9,15]:=1616302937;
   	OWF_Key[9,16]:=182946603;
   	OWF_Key[10,13]:=1325878573;
   	OWF_Key[10,14]:=1945679484;
   	OWF_Key[10,15]:=198793809;
   	OWF_Key[10,16]:=1919335442;
   	OWF_Key[11,13]:=1564455476;
   	OWF_Key[11,14]:=643845182;
   	OWF_Key[11,15]:=1627849411;
   	OWF_Key[11,16]:=1185245357;
   	OWF_Key[12,13]:=1917947303;
   	OWF_Key[12,14]:=561134487;
   	OWF_Key[12,15]:=453014383;
   	OWF_Key[12,16]:=290220751;
   	OWF_Key[13,13]:=1258679728;
   	OWF_Key[13,14]:=649968820;
   	OWF_Key[13,15]:=809905849;
   	OWF_Key[13,16]:=560836421;
   	OWF_Key[14,13]:=482755903;
   	OWF_Key[14,14]:=919140814;
   	OWF_Key[14,15]:=979596316;
   	OWF_Key[14,16]:=1735062741;
   	OWF_Key[15,13]:=1362928281;
   	OWF_Key[15,14]:=2061487261;
   	OWF_Key[15,15]:=285408975;
   	OWF_Key[15,16]:=180370867;
   	OWF_Key[16,13]:=670546063;
   	OWF_Key[16,14]:=712104113;
   	OWF_Key[16,15]:=1951589450;
   	OWF_Key[16,16]:=1738253114;
   	OWF_Key[17,13]:=1669460550;
   	OWF_Key[17,14]:=1403355642;
   	OWF_Key[17,15]:=1129897394;
   	OWF_Key[17,16]:=1783591382;
   	OWF_Key[18,13]:=1064160739;
   	OWF_Key[18,14]:=888090837;
   	OWF_Key[18,15]:=1910618387;
   	OWF_Key[18,16]:=1458664956;
   	OWF_Key[19,13]:=1151080277;
   	OWF_Key[19,14]:=420116810;
   	OWF_Key[19,15]:=1893442335;
   	OWF_Key[19,16]:=1425027207;
   	OWF_Key[20,13]:=428816941;
   	OWF_Key[20,14]:=1662558165;
   	OWF_Key[20,15]:=307375973;
   	OWF_Key[20,16]:=533927155;
   	OWF_Key[21,13]:=1264084049;
   	OWF_Key[21,14]:=1926233168;
   	OWF_Key[21,15]:=525930072;
   	OWF_Key[21,16]:=1719696135;
   	OWF_Key[22,13]:=978289204;
   	OWF_Key[22,14]:=379512271;
   	OWF_Key[22,15]:=1026840126;
   	OWF_Key[22,16]:=765316908;
   	OWF_Key[23,13]:=901692748;
   	OWF_Key[23,14]:=1577626792;
   	OWF_Key[23,15]:=547638324;
   	OWF_Key[23,16]:=252696951;
   	OWF_Key[24,13]:=1490534977;
   	OWF_Key[24,14]:=1821556895;
   	OWF_Key[24,15]:=2092883059;
   	OWF_Key[24,16]:=1739124451;
   	OWF_Key[25,13]:=886462231;
   	OWF_Key[25,14]:=1842653560;
   	OWF_Key[25,15]:=1093841042;
   	OWF_Key[25,16]:=457940159;
   	OWF_Key[26,13]:=902257555;
   	OWF_Key[26,14]:=1094025454;
   	OWF_Key[26,15]:=134405645;
   	OWF_Key[26,16]:=41176787;
   	OWF_Key[27,13]:=412607945;
   	OWF_Key[27,14]:=1952067299;
   	OWF_Key[27,15]:=353747084;
   	OWF_Key[27,16]:=1682000323;
   	OWF_Key[28,13]:=18005791;
   	OWF_Key[28,14]:=620821249;
   	OWF_Key[28,15]:=1113212535;
   	OWF_Key[28,16]:=897987427;
   	OWF_Key[29,13]:=1190050746;
   	OWF_Key[29,14]:=643899149;
   	OWF_Key[29,15]:=722485001;
   	OWF_Key[29,16]:=893986043;
   	OWF_Key[30,13]:=1098154477;
   	OWF_Key[30,14]:=1637361182;
   	OWF_Key[30,15]:=978110562;
   	OWF_Key[30,16]:=550604029;
   	OWF_Key[31,13]:=592959310;
   	OWF_Key[31,14]:=978865608;
   	OWF_Key[31,15]:=1198404585;
   	OWF_Key[31,16]:=419804619;
   	OWF_Key[32,13]:=145480636;
   	OWF_Key[32,14]:=626472266;
   	OWF_Key[32,15]:=1453538134;